FUNCTION_BLOCK "X_Simulacia"   // FB100, LAD
{ S7_Optimized_Access := 'TRUE' }
VERSION : 0.1
   VAR
      Servis : Struct
         Bag : Bool;
         BoxSmall : Bool;
         BoxLarge : Bool;
         Con_Printer : Bool;
      END_STRUCT;
      BagServis : String;
      BoxServis : String;
      OPC_Con : Struct
         NewMDR_Flag : String;
         NewArticleFlag : String;
         NewBatchNumber : String;
         NewArtBaseNumber : DInt;
         NewMarketREG_Code : String;
         NewBatchEndTime : String;
         NewExtDate : String;
      END_STRUCT;
      Artikel1 : Struct
         bag_dmc_code : Array[0..9] of Char;
         box_dmc_code : Array[0..9] of Char;
      END_STRUCT;
      Artikel2 : Struct
         bag_dmc_code : Array[0..9] of Char;
         box_dmc_code : Array[0..9] of Char;
      END_STRUCT;
      Artikel3 : Struct
         bag_dmc_code : Array[0..9] of Char;
         box_dmc_code : Array[0..9] of Char;
      END_STRUCT;
      TRP_Materia : "UDT_TRP_Comm";
      Artikel4 : Struct
         bag_dmc_code : Array[0..9] of Char;
         box_dmc_code : Array[0..9] of Char;
      END_STRUCT;
   END_VAR
   VAR RETAIN
      IEC_Counter_0_Instance : CTU_INT;
      Count : Int;
   END_VAR
   VAR
      ResetCount : Bool;
      Log0 : Bool;
      Log1 : Bool;
      bag_dmc_code : Array[0..9] of Char;
      box_dmc_code : Array[0..9] of Char;
      article_num : Array[0..11] of Char;
      total_in_bag : Array[0..6] of Char;
      total_in_box : Array[0..6] of Char;
      product_weight : Array[0..9] of Char;
      line_number : Array[0..4] of Char;
      order_num : Array[0..11] of Char;
   END_VAR
   VAR_TEMP
      TmpI : Int;
      TmpD : DInt;
      TmpU : UInt;
   END_VAR
   // Artikel1.bag_dmc_code[0] := '0';
   // Artikel1.bag_dmc_code[1] := '0';
   // Artikel1.bag_dmc_code[2] := '0';
   // Artikel1.bag_dmc_code[3] := '4';
   // Artikel1.bag_dmc_code[4] := '6';
   // Artikel1.bag_dmc_code[5] := '0';
   // Artikel1.bag_dmc_code[6] := '3';
   // Artikel1.bag_dmc_code[7] := '6';
   // Artikel1.bag_dmc_code[8] := '4';
   // Artikel1.bag_dmc_code[9] := '3';
   // Artikel1.box_dmc_code[9] := '3';
   // Artikel1.box_dmc_code[8] := '2';
   // Artikel1.box_dmc_code[7] := '2';
   // Artikel1.box_dmc_code[6] := '7';
   // Artikel1.box_dmc_code[5] := '4';
   // Artikel1.box_dmc_code[4] := '6';
   // Artikel1.box_dmc_code[3] := '4';
   // Artikel1.box_dmc_code[2] := '0';
   // Artikel1.box_dmc_code[1] := '0';
   // Artikel1.box_dmc_code[0] := '0';
   // TRP_Materia.NewMachineID := '999';
   // TRP_Materia.NewArticleNumber := 76166100;
   // TRP_Materia.NewBatchNumber := '1011234580';
   // TRP_Materia.NewGTIN_Number := '07322541067896';
   // article_num[0] := '$04';
   // article_num[1] := '$05';
   // article_num[2] := '$06';
   // article_num[3] := '$07';
   // article_num[4] := '$08';
   // article_num[5] := '$04';
   // article_num[6] := '$05';
   // article_num[7] := '$06';
   // article_num[8] := '$05';
   // article_num[9] := '$03';
   // article_num[10] := '$02';
   // article_num[11] := '$01';
   // order_num[0] := '$03';
   // order_num[1] := '$03';
   // order_num[2] := '$03';
   // Artikel2.bag_dmc_code[0] := '0';
   // Artikel2.bag_dmc_code[9] := '2';
   // Artikel2.bag_dmc_code[8] := '3';
   // Artikel2.bag_dmc_code[7] := '6';
   // Artikel2.bag_dmc_code[6] := '7';
   // Artikel2.bag_dmc_code[5] := '7';
   // Artikel2.bag_dmc_code[4] := '6';
   // Artikel2.bag_dmc_code[3] := '3';
   // Artikel2.bag_dmc_code[2] := '0';
   // Artikel2.bag_dmc_code[1] := '0';
BEGIN

REGION Network 1
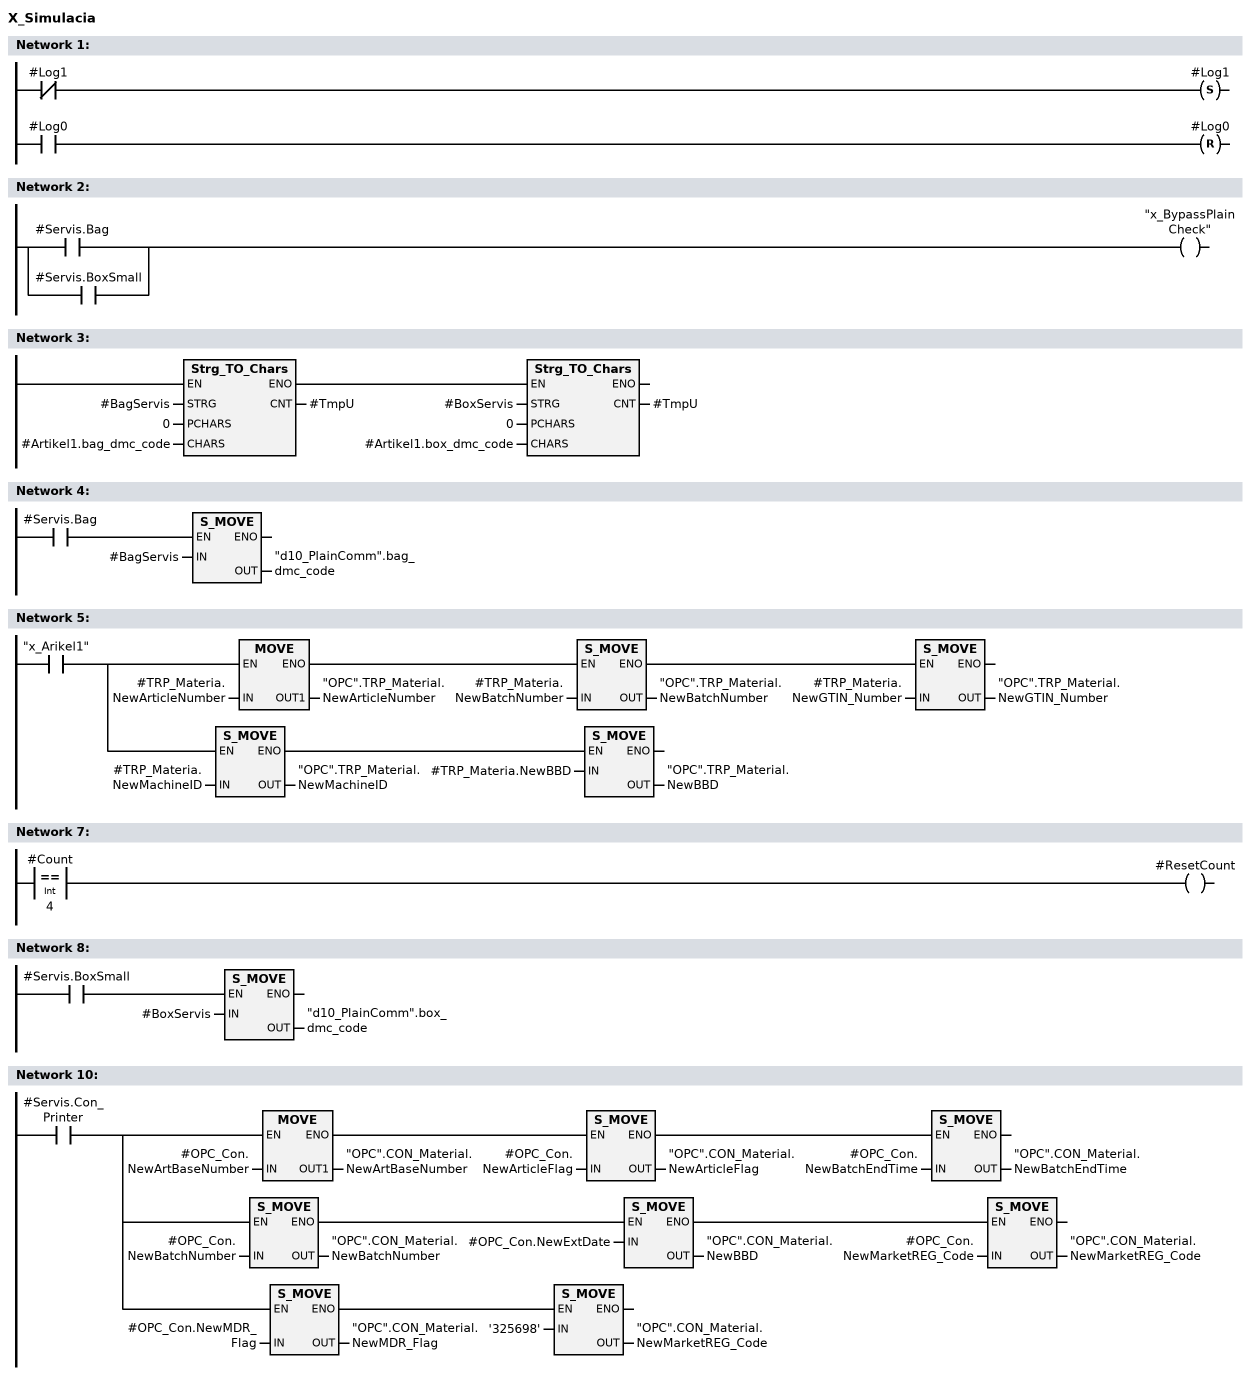
   RUNG wire#powerrail
      I_Contact( #Log1 )
      S_Coil( #Log1 )
   END_RUNG
   RUNG wire#powerrail
      Contact( #Log0 )
      R_Coil( #Log0 )
   END_RUNG
   // the same network as SCL:
   IF NOT #Log1 THEN #Log1 := TRUE; END_IF;
   IF #Log0 THEN #Log0 := FALSE; END_IF;
END_REGION

REGION Network 2
   RUNG wire#powerrail
      Contact( #Servis.Bag )
      wire#w1
      Coil( "x_BypassPlainCheck" )
   END_RUNG
   RUNG wire#powerrail
      Contact( #Servis.BoxSmall )
   END_RUNG wire#w1
   // the same network as SCL:
   "x_BypassPlainCheck" := #Servis.Bag OR #Servis.BoxSmall;
END_REGION

REGION Network 3
   // no SCL statement known for Strg_TO_Chars: written as a call
   // ENO of a box is taken as its EN; it also drops when the box reports an error
   Strg_TO_Chars(Strg := #BagServis, pChars := 0, Chars := #Artikel1.bag_dmc_code, Cnt => #TmpU);
   Strg_TO_Chars(Strg := #BoxServis, pChars := 0, Chars := #Artikel1.box_dmc_code, Cnt => #TmpU);
END_REGION

REGION Network 4
   RUNG wire#powerrail
      Contact( #Servis.Bag )
      S_Move(in := #BagServis, out => "d10_PlainComm".bag_dmc_code)
   END_RUNG
   // the same network as SCL:
   IF #Servis.Bag THEN "d10_PlainComm".bag_dmc_code := #BagServis; END_IF;
END_REGION

REGION Network 5
   RUNG wire#powerrail
      Contact( "x_Arikel1" )
      wire#w1
      Move(in := #TRP_Materia.NewArticleNumber, out1 => "OPC".TRP_Material.NewArticleNumber)
      S_Move(in := #TRP_Materia.NewBatchNumber, out => "OPC".TRP_Material.NewBatchNumber)
      S_Move(in := #TRP_Materia.NewGTIN_Number, out => "OPC".TRP_Material.NewGTIN_Number)
   END_RUNG
   RUNG wire#w1
      S_Move(in := #TRP_Materia.NewMachineID, out => "OPC".TRP_Material.NewMachineID)
      S_Move(in := #TRP_Materia.NewBBD, out => "OPC".TRP_Material.NewBBD)
   END_RUNG
   // the same network as SCL:
   IF "x_Arikel1" THEN
       "OPC".TRP_Material.NewArticleNumber := #TRP_Materia.NewArticleNumber;
       "OPC".TRP_Material.NewBatchNumber := #TRP_Materia.NewBatchNumber;
       "OPC".TRP_Material.NewGTIN_Number := #TRP_Materia.NewGTIN_Number;
       "OPC".TRP_Material.NewMachineID := #TRP_Materia.NewMachineID;
       "OPC".TRP_Material.NewBBD := #TRP_Materia.NewBBD;
   END_IF;
END_REGION

REGION Network 7
   RUNG wire#powerrail
      { S7_Templates := "SrcType := Int" } EQ_Contact(in1 := #Count, in2 := 4)
      Coil( #ResetCount )
   END_RUNG
   // the same network as SCL:
   #ResetCount := #Count = 4;
END_REGION

REGION Network 8
   RUNG wire#powerrail
      Contact( #Servis.BoxSmall )
      S_Move(in := #BoxServis, out => "d10_PlainComm".box_dmc_code)
   END_RUNG
   // the same network as SCL:
   IF #Servis.BoxSmall THEN "d10_PlainComm".box_dmc_code := #BoxServis; END_IF;
END_REGION

REGION Network 10
   RUNG wire#powerrail
      Contact( #Servis.Con_Printer )
      wire#w1
      Move(in := #OPC_Con.NewArtBaseNumber, out1 => "OPC".CON_Material.NewArtBaseNumber)
      S_Move(in := #OPC_Con.NewArticleFlag, out => "OPC".CON_Material.NewArticleFlag)
      S_Move(in := #OPC_Con.NewBatchEndTime, out => "OPC".CON_Material.NewBatchEndTime)
   END_RUNG
   RUNG wire#w1
      S_Move(in := #OPC_Con.NewBatchNumber, out => "OPC".CON_Material.NewBatchNumber)
      S_Move(in := #OPC_Con.NewExtDate, out => "OPC".CON_Material.NewBBD)
      S_Move(in := #OPC_Con.NewMarketREG_Code, out => "OPC".CON_Material.NewMarketREG_Code)
   END_RUNG
   RUNG wire#w1
      S_Move(in := #OPC_Con.NewMDR_Flag, out => "OPC".CON_Material.NewMDR_Flag)
      S_Move(in := '325698', out => "OPC".CON_Material.NewMarketREG_Code)
   END_RUNG
   // the same network as SCL:
   IF #Servis.Con_Printer THEN
       "OPC".CON_Material.NewArtBaseNumber := #OPC_Con.NewArtBaseNumber;
       "OPC".CON_Material.NewArticleFlag := #OPC_Con.NewArticleFlag;
       "OPC".CON_Material.NewBatchEndTime := #OPC_Con.NewBatchEndTime;
       "OPC".CON_Material.NewBatchNumber := #OPC_Con.NewBatchNumber;
       "OPC".CON_Material.NewBBD := #OPC_Con.NewExtDate;
       "OPC".CON_Material.NewMarketREG_Code := #OPC_Con.NewMarketREG_Code;
       "OPC".CON_Material.NewMDR_Flag := #OPC_Con.NewMDR_Flag;
       "OPC".CON_Material.NewMarketREG_Code := '325698';
   END_IF;
END_REGION
END_FUNCTION_BLOCK

FUNCTION_BLOCK "DMCC"   // FB102, LAD
{ S7_Optimized_Access := 'TRUE' }
VERSION : 0.1
   VAR_INPUT
      Reset_Camera_Box : Bool;
      Set_Camera_Box : Bool;
      Reboot : Bool;
      Reset : Bool;
      FPS_Camera_Box : Int;
   END_VAR
   VAR_OUTPUT
      Lenght_Camera_Box : Int;
      Execute_Camera_Box : Bool;
      Error : Bool;
   END_VAR
   VAR
      Edge : Array[0..15] of Bool;
      Camera_Box : Struct
         NumberFPS : String;
         ClearBufferR : Bool;
         ClearBufferR2 : Bool;
         ClearLogR : Bool;
         ClearLogR2 : Bool;
         Log : Bool;
         RequestReset : Bool;
         RequestSet : Bool;
         RebootRequest : Bool;
         RebootE : Bool;
         SetS : String;
      END_STRUCT;
      log0 : Bool;
      t_Error : TON_TIME;
      t_Error2 : TON_TIME;
   END_VAR
   VAR_TEMP
      TmpUInt : UInt;
      TmpI : Int;
      TmpS : String;
      TmpS2 : String;
   END_VAR
   VAR CONSTANT
      ResetBuffer : String := '||>COM.BUFFER-RESET';
      ClerarDeviceLog : String := '||>DEVICE-LOG.CLEAR';
      SetCameraS : String := '||>SET CAMERA.BURST-LENGTH ';
      SetCameraS_bag : String := '||>SET CAMERA.BURST-LENGTH ';
      RebootS : String := '||>REBOOT';
   END_VAR
   VAR_TEMP   // added for the SCL form of the ladder/FBD networks
      _w1 : Bool;
      _w2 : Bool;
      _w3 : Bool;
   END_VAR
BEGIN

REGION Network 1
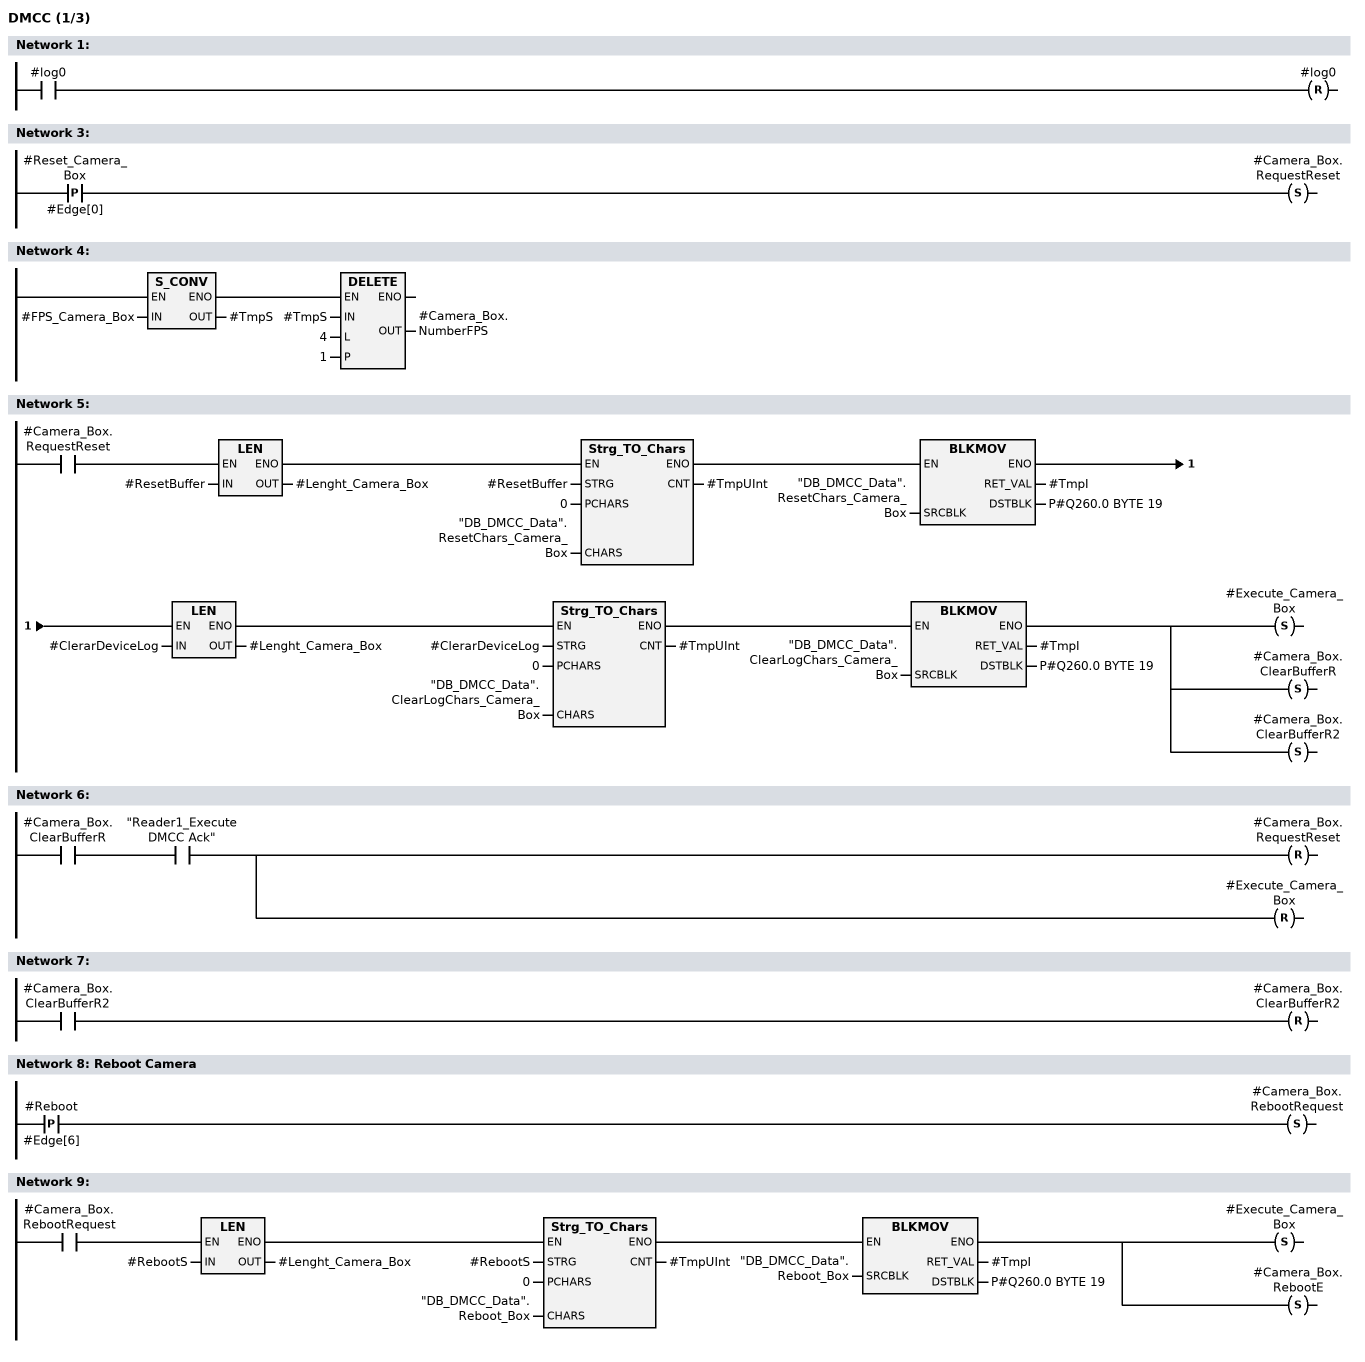
   RUNG wire#powerrail
      Contact( #log0 )
      R_Coil( #log0 )
   END_RUNG
   // the same network as SCL:
   IF #log0 THEN #log0 := FALSE; END_IF;
END_REGION

REGION Network 3
   RUNG wire#powerrail
      P_Contact(operand := #Reset_Camera_Box, bit := #Edge[0])
      S_Coil( #Camera_Box.RequestReset )
   END_RUNG
   // the same network as SCL:
   #_w1 := #Reset_Camera_Box AND NOT #Edge[0];   // rising edge of #Reset_Camera_Box
   #Edge[0] := #Reset_Camera_Box;
   IF #_w1 THEN #Camera_Box.RequestReset := TRUE; END_IF;
END_REGION

REGION Network 4
   #TmpS := S_CONV(IN := #FPS_Camera_Box);
   #Camera_Box.NumberFPS := DELETE(IN := #TmpS, L := 4, P := 1);
END_REGION

REGION Network 5
   // no SCL statement known for Strg_TO_Chars: written as a call
   // ENO of a box is taken as its EN; it also drops when the box reports an error
   IF #Camera_Box.RequestReset THEN
       #Lenght_Camera_Box := LEN(IN := #ResetBuffer);
       Strg_TO_Chars(Strg := #ResetBuffer,
                     pChars := 0,
                     Chars := "DB_DMCC_Data".ResetChars_Camera_Box,
                     Cnt => #TmpUInt);
       #TmpI := BLKMOV(SRCBLK := "DB_DMCC_Data".ResetChars_Camera_Box, DSTBLK => P#Q260.0 BYTE 19);
       #Lenght_Camera_Box := LEN(IN := #ClerarDeviceLog);
       Strg_TO_Chars(Strg := #ClerarDeviceLog,
                     pChars := 0,
                     Chars := "DB_DMCC_Data".ClearLogChars_Camera_Box,
                     Cnt => #TmpUInt);
       #TmpI := BLKMOV(SRCBLK := "DB_DMCC_Data".ClearLogChars_Camera_Box, DSTBLK => P#Q260.0 BYTE 19);
       #Execute_Camera_Box := TRUE;
       #Camera_Box.ClearBufferR := TRUE;
       #Camera_Box.ClearBufferR2 := TRUE;
   END_IF;
END_REGION

REGION Network 6
   RUNG wire#powerrail
      Contact( #Camera_Box.ClearBufferR )
      Contact( "Reader1_Execute DMCC Ack" )
      wire#w1
      R_Coil( #Camera_Box.RequestReset )
   END_RUNG
   RUNG wire#w1
      R_Coil( #Execute_Camera_Box )
   END_RUNG
   // the same network as SCL:
   IF #Camera_Box.ClearBufferR AND "Reader1_Execute DMCC Ack" THEN
       #Camera_Box.RequestReset := FALSE;
       #Execute_Camera_Box := FALSE;
   END_IF;
END_REGION

REGION Network 7
   RUNG wire#powerrail
      Contact( #Camera_Box.ClearBufferR2 )
      R_Coil( #Camera_Box.ClearBufferR2 )
   END_RUNG
   // the same network as SCL:
   IF #Camera_Box.ClearBufferR2 THEN #Camera_Box.ClearBufferR2 := FALSE; END_IF;
END_REGION

REGION Network 8: Reboot Camera
   RUNG wire#powerrail
      P_Contact(operand := #Reboot, bit := #Edge[6])
      S_Coil( #Camera_Box.RebootRequest )
   END_RUNG
   // the same network as SCL:
   #_w1 := #Reboot AND NOT #Edge[6];   // rising edge of #Reboot
   #Edge[6] := #Reboot;
   IF #_w1 THEN #Camera_Box.RebootRequest := TRUE; END_IF;
END_REGION

REGION Network 9
   // no SCL statement known for Strg_TO_Chars: written as a call
   // ENO of a box is taken as its EN; it also drops when the box reports an error
   IF #Camera_Box.RebootRequest THEN
       #Lenght_Camera_Box := LEN(IN := #RebootS);
       Strg_TO_Chars(Strg := #RebootS, pChars := 0, Chars := "DB_DMCC_Data".Reboot_Box, Cnt => #TmpUInt);
       #TmpI := BLKMOV(SRCBLK := "DB_DMCC_Data".Reboot_Box, DSTBLK => P#Q260.0 BYTE 19);
       #Execute_Camera_Box := TRUE;
       #Camera_Box.RebootE := TRUE;
   END_IF;
END_REGION

REGION Network 10
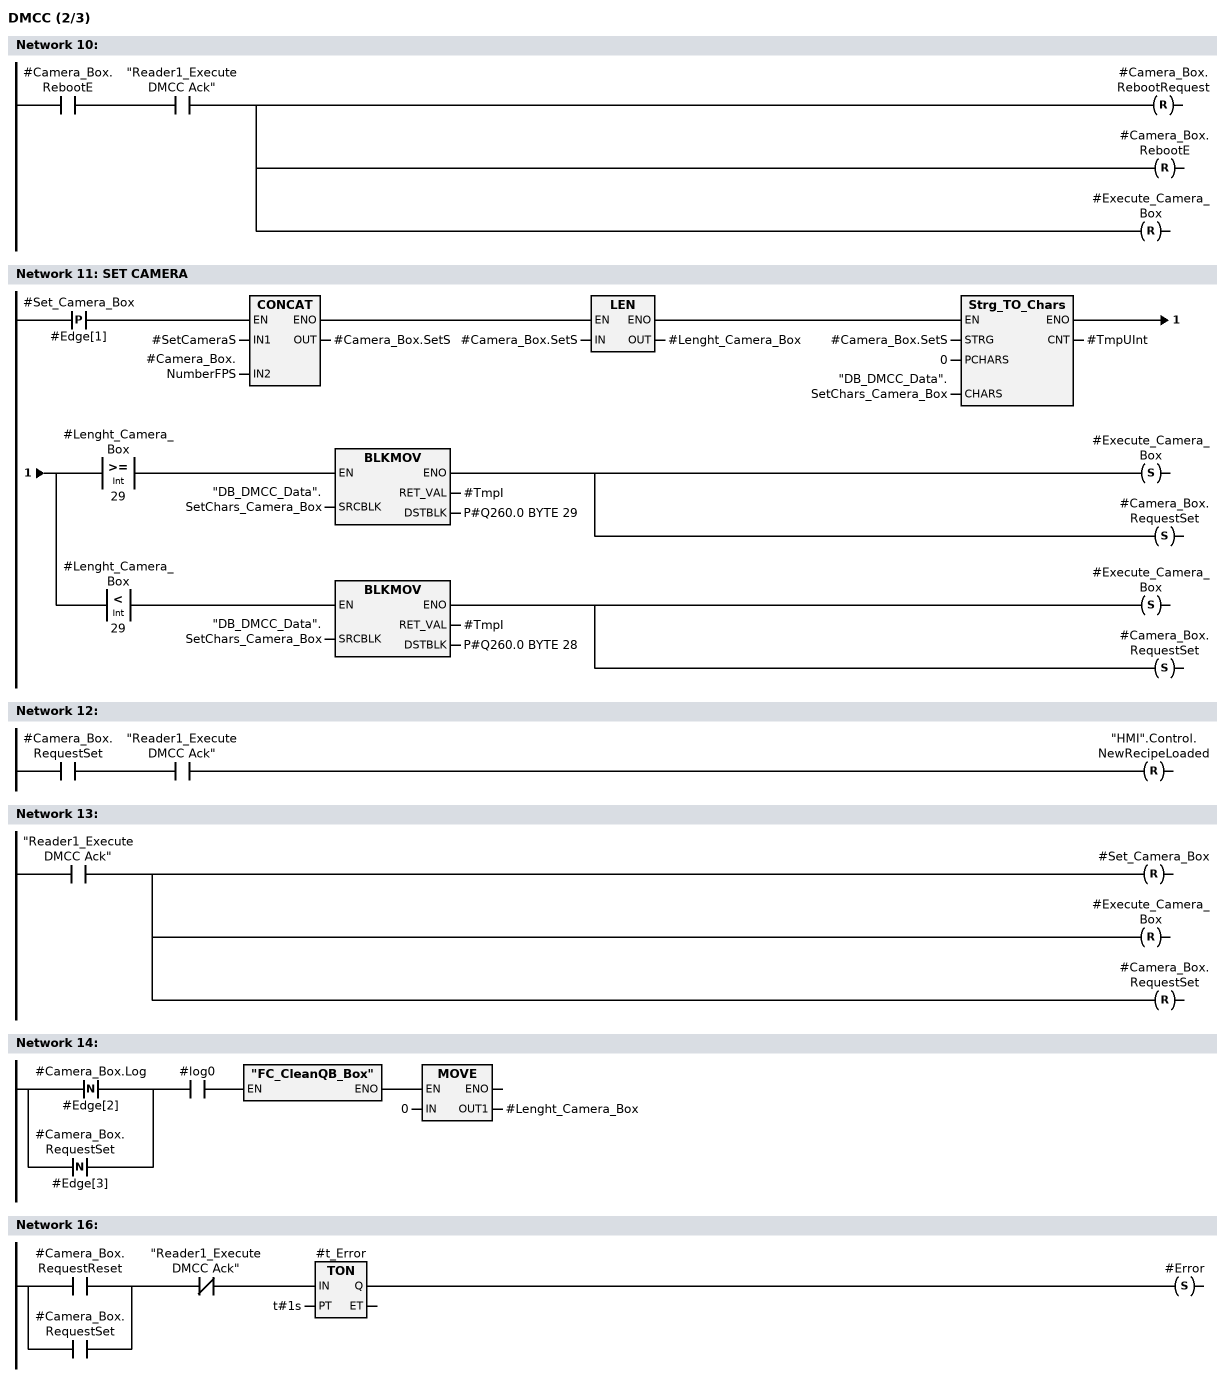
   RUNG wire#powerrail
      Contact( #Camera_Box.RebootE )
      Contact( "Reader1_Execute DMCC Ack" )
      wire#w1
      R_Coil( #Camera_Box.RebootRequest )
   END_RUNG
   RUNG wire#w1
      R_Coil( #Camera_Box.RebootE )
   END_RUNG
   RUNG wire#w1
      R_Coil( #Execute_Camera_Box )
   END_RUNG
   // the same network as SCL:
   IF #Camera_Box.RebootE AND "Reader1_Execute DMCC Ack" THEN #Camera_Box.RebootRequest := FALSE; END_IF;
   #_w1 := #Camera_Box.RebootE AND "Reader1_Execute DMCC Ack";
   IF #_w1 THEN
       #Camera_Box.RebootE := FALSE;
       #Execute_Camera_Box := FALSE;
   END_IF;
END_REGION

REGION Network 11: SET CAMERA
   // no SCL statement known for Strg_TO_Chars: written as a call
   // ENO of a box is taken as its EN; it also drops when the box reports an error
   #_w1 := #Set_Camera_Box AND NOT #Edge[1];   // rising edge of #Set_Camera_Box
   #Edge[1] := #Set_Camera_Box;
   IF #_w1 THEN
       #Camera_Box.SetS := CONCAT(IN1 := #SetCameraS, IN2 := #Camera_Box.NumberFPS);
       #Lenght_Camera_Box := LEN(IN := #Camera_Box.SetS);
       Strg_TO_Chars(Strg := #Camera_Box.SetS,
                     pChars := 0,
                     Chars := "DB_DMCC_Data".SetChars_Camera_Box,
                     Cnt => #TmpUInt);
   END_IF;
   IF #_w1 AND (#Lenght_Camera_Box >= 29) THEN
       #TmpI := BLKMOV(SRCBLK := "DB_DMCC_Data".SetChars_Camera_Box, DSTBLK => P#Q260.0 BYTE 29);
       #Execute_Camera_Box := TRUE;
       #Camera_Box.RequestSet := TRUE;
   END_IF;
   IF #_w1 AND (#Lenght_Camera_Box < 29) THEN
       #TmpI := BLKMOV(SRCBLK := "DB_DMCC_Data".SetChars_Camera_Box, DSTBLK => P#Q260.0 BYTE 28);
       #Execute_Camera_Box := TRUE;
       #Camera_Box.RequestSet := TRUE;
   END_IF;
END_REGION

REGION Network 12
   RUNG wire#powerrail
      Contact( #Camera_Box.RequestSet )
      Contact( "Reader1_Execute DMCC Ack" )
      R_Coil( "HMI".Control.NewRecipeLoaded )
   END_RUNG
   // the same network as SCL:
   IF #Camera_Box.RequestSet AND "Reader1_Execute DMCC Ack" THEN
       "HMI".Control.NewRecipeLoaded := FALSE;
   END_IF;
END_REGION

REGION Network 13
   RUNG wire#powerrail
      Contact( "Reader1_Execute DMCC Ack" )
      wire#w1
      R_Coil( #Set_Camera_Box )
   END_RUNG
   RUNG wire#w1
      R_Coil( #Execute_Camera_Box )
   END_RUNG
   RUNG wire#w1
      R_Coil( #Camera_Box.RequestSet )
   END_RUNG
   // the same network as SCL:
   IF "Reader1_Execute DMCC Ack" THEN
       #Set_Camera_Box := FALSE;
       #Execute_Camera_Box := FALSE;
       #Camera_Box.RequestSet := FALSE;
   END_IF;
END_REGION

REGION Network 14
   RUNG wire#powerrail
      N_Contact(operand := #Camera_Box.Log, bit := #Edge[2])
      wire#w1
      Contact( #log0 )
      "FC_CleanQB_Box"()
      Move(in := 0, out1 => #Lenght_Camera_Box)
   END_RUNG
   RUNG wire#powerrail
      N_Contact(operand := #Camera_Box.RequestSet, bit := #Edge[3])
   END_RUNG wire#w1
   // the same network as SCL:
   #_w1 := NOT #Camera_Box.Log AND #Edge[2];   // falling edge of #Camera_Box.Log
   #Edge[2] := #Camera_Box.Log;
   #_w2 := NOT #Camera_Box.RequestSet AND #Edge[3];   // falling edge of #Camera_Box.RequestSet
   #Edge[3] := #Camera_Box.RequestSet;
   "FC_CleanQB_Box"(EN := (#_w1 OR #_w2) AND #log0, ENO => #_w3);
   IF #_w3 THEN #Lenght_Camera_Box := 0; END_IF;
END_REGION

REGION Network 16
   #t_Error(IN := (#Camera_Box.RequestReset OR #Camera_Box.RequestSet) AND NOT "Reader1_Execute DMCC Ack",   // TON
            PT := t#1s);
   IF #t_Error.Q THEN #Error := TRUE; END_IF;
END_REGION

REGION Network 17
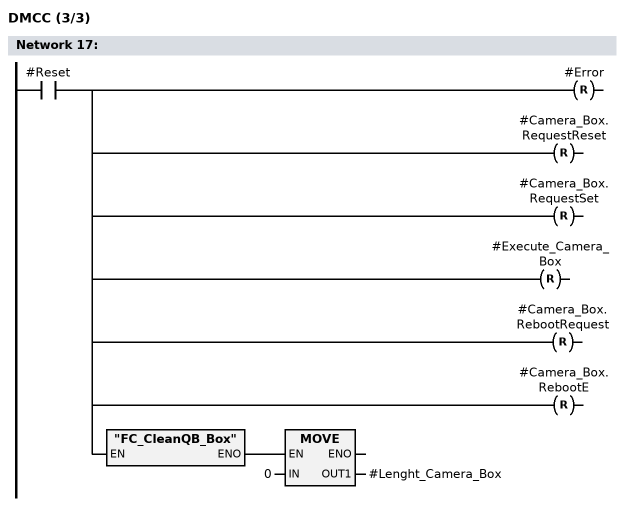
   RUNG wire#powerrail
      Contact( #Reset )
      wire#w1
      R_Coil( #Error )
   END_RUNG
   RUNG wire#w1
      R_Coil( #Camera_Box.RequestReset )
   END_RUNG
   RUNG wire#w1
      R_Coil( #Camera_Box.RequestSet )
   END_RUNG
   RUNG wire#w1
      R_Coil( #Execute_Camera_Box )
   END_RUNG
   RUNG wire#w1
      R_Coil( #Camera_Box.RebootRequest )
   END_RUNG
   RUNG wire#w1
      R_Coil( #Camera_Box.RebootE )
   END_RUNG
   RUNG wire#w1
      "FC_CleanQB_Box"()
      Move(in := 0, out1 => #Lenght_Camera_Box)
   END_RUNG
   // the same network as SCL:
   IF #Reset THEN
       #Error := FALSE;
       #Camera_Box.RequestReset := FALSE;
       #Camera_Box.RequestSet := FALSE;
       #Execute_Camera_Box := FALSE;
       #Camera_Box.RebootRequest := FALSE;
       #Camera_Box.RebootE := FALSE;
   END_IF;
   "FC_CleanQB_Box"(EN := #Reset, ENO => #_w1);
   IF #_w1 THEN #Lenght_Camera_Box := 0; END_IF;
END_REGION
END_FUNCTION_BLOCK

FUNCTION_BLOCK "DMCC_bag"   // FB103, LAD
{ S7_Optimized_Access := 'TRUE' }
VERSION : 0.1
   VAR_INPUT
      Reset_Camera_Bag : Bool;
      Set_Camera_Bag : Bool;
      Reset : Bool;
      Reboot : Bool;
      FPS_Camera_Boag : Int;
   END_VAR
   VAR_OUTPUT
      Lenght_Camera_Bag : Int;
      Execute_Camera_Bag : Bool;
      Error : Bool;
   END_VAR
   VAR
      Edge : Array[0..15] of Bool;
      Camera_Bag : Struct
         NumberFPS : String;
         ClearBufferR : Bool;
         ClearBufferR2 : Bool;
         ClearLogR : Bool;
         ClearLogR2 : Bool;
         Log : Bool;
         RequestReset : Bool;
         RequestSet : Bool;
         RebootRequest : Bool;
         RebootE : Bool;
         SetS : String;
      END_STRUCT;
      log0 : Bool;
      t_Error : TON_TIME;
      t_Error2 : TON_TIME;
   END_VAR
   VAR_TEMP
      TmpUInt : UInt;
      TmpI : Int;
      TmpS : String;
      TmpS2 : String;
   END_VAR
   VAR CONSTANT
      ResetBuffer : String := '||>COM.BUFFER-RESET';
      ClerarDeviceLog : String := '||>DEVICE-LOG.CLEAR';
      SetCameraS : String := '||>SET CAMERA.BURST-LENGTH ';
      RebootS : String := '||>REBOOT';
   END_VAR
   VAR_TEMP   // added for the SCL form of the ladder/FBD networks
      _w1 : Bool;
      _w2 : Bool;
      _w3 : Bool;
   END_VAR
BEGIN

REGION Network 2
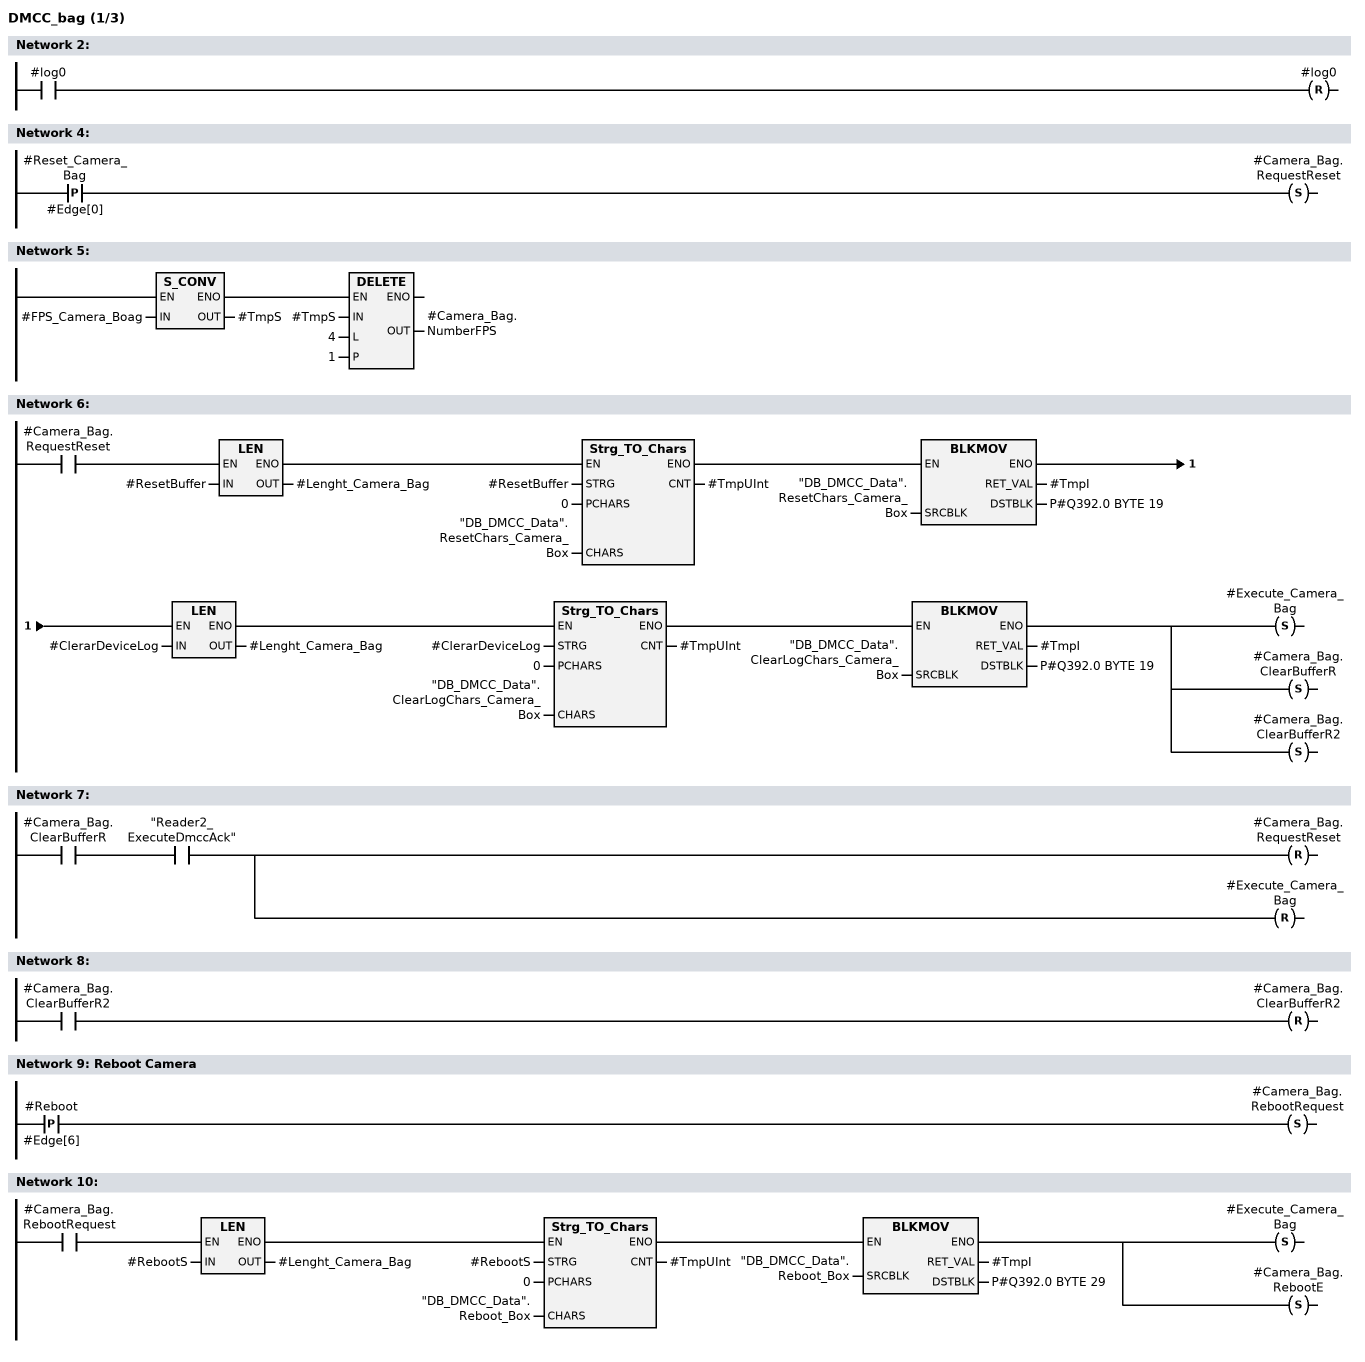
   RUNG wire#powerrail
      Contact( #log0 )
      R_Coil( #log0 )
   END_RUNG
   // the same network as SCL:
   IF #log0 THEN #log0 := FALSE; END_IF;
END_REGION

REGION Network 4
   RUNG wire#powerrail
      P_Contact(operand := #Reset_Camera_Bag, bit := #Edge[0])
      S_Coil( #Camera_Bag.RequestReset )
   END_RUNG
   // the same network as SCL:
   #_w1 := #Reset_Camera_Bag AND NOT #Edge[0];   // rising edge of #Reset_Camera_Bag
   #Edge[0] := #Reset_Camera_Bag;
   IF #_w1 THEN #Camera_Bag.RequestReset := TRUE; END_IF;
END_REGION

REGION Network 5
   #TmpS := S_CONV(IN := #FPS_Camera_Boag);
   #Camera_Bag.NumberFPS := DELETE(IN := #TmpS, L := 4, P := 1);
END_REGION

REGION Network 6
   // no SCL statement known for Strg_TO_Chars: written as a call
   // ENO of a box is taken as its EN; it also drops when the box reports an error
   IF #Camera_Bag.RequestReset THEN
       #Lenght_Camera_Bag := LEN(IN := #ResetBuffer);
       Strg_TO_Chars(Strg := #ResetBuffer,
                     pChars := 0,
                     Chars := "DB_DMCC_Data".ResetChars_Camera_Box,
                     Cnt => #TmpUInt);
       #TmpI := BLKMOV(SRCBLK := "DB_DMCC_Data".ResetChars_Camera_Box, DSTBLK => P#Q392.0 BYTE 19);
       #Lenght_Camera_Bag := LEN(IN := #ClerarDeviceLog);
       Strg_TO_Chars(Strg := #ClerarDeviceLog,
                     pChars := 0,
                     Chars := "DB_DMCC_Data".ClearLogChars_Camera_Box,
                     Cnt => #TmpUInt);
       #TmpI := BLKMOV(SRCBLK := "DB_DMCC_Data".ClearLogChars_Camera_Box, DSTBLK => P#Q392.0 BYTE 19);
       #Execute_Camera_Bag := TRUE;
       #Camera_Bag.ClearBufferR := TRUE;
       #Camera_Bag.ClearBufferR2 := TRUE;
   END_IF;
END_REGION

REGION Network 7
   RUNG wire#powerrail
      Contact( #Camera_Bag.ClearBufferR )
      Contact( "Reader2_ExecuteDmccAck" )
      wire#w1
      R_Coil( #Camera_Bag.RequestReset )
   END_RUNG
   RUNG wire#w1
      R_Coil( #Execute_Camera_Bag )
   END_RUNG
   // the same network as SCL:
   IF #Camera_Bag.ClearBufferR AND "Reader2_ExecuteDmccAck" THEN
       #Camera_Bag.RequestReset := FALSE;
       #Execute_Camera_Bag := FALSE;
   END_IF;
END_REGION

REGION Network 8
   RUNG wire#powerrail
      Contact( #Camera_Bag.ClearBufferR2 )
      R_Coil( #Camera_Bag.ClearBufferR2 )
   END_RUNG
   // the same network as SCL:
   IF #Camera_Bag.ClearBufferR2 THEN #Camera_Bag.ClearBufferR2 := FALSE; END_IF;
END_REGION

REGION Network 9: Reboot Camera
   RUNG wire#powerrail
      P_Contact(operand := #Reboot, bit := #Edge[6])
      S_Coil( #Camera_Bag.RebootRequest )
   END_RUNG
   // the same network as SCL:
   #_w1 := #Reboot AND NOT #Edge[6];   // rising edge of #Reboot
   #Edge[6] := #Reboot;
   IF #_w1 THEN #Camera_Bag.RebootRequest := TRUE; END_IF;
END_REGION

REGION Network 10
   // no SCL statement known for Strg_TO_Chars: written as a call
   // ENO of a box is taken as its EN; it also drops when the box reports an error
   IF #Camera_Bag.RebootRequest THEN
       #Lenght_Camera_Bag := LEN(IN := #RebootS);
       Strg_TO_Chars(Strg := #RebootS, pChars := 0, Chars := "DB_DMCC_Data".Reboot_Box, Cnt => #TmpUInt);
       #TmpI := BLKMOV(SRCBLK := "DB_DMCC_Data".Reboot_Box, DSTBLK => P#Q392.0 BYTE 29);
       #Execute_Camera_Bag := TRUE;
       #Camera_Bag.RebootE := TRUE;
   END_IF;
END_REGION

REGION Network 11